// Mitsubishi GX Works2 project: 11国轩烘烤线体修改1028   PLC: Q06UDEH

TYPE ConveyorIO : STRUCT
  xUnloadCCW : BOOL;  (* 下料为反转 *)
  xUnloadAlarm : BOOL;  (* 下料报警 *)
  xUnload : BOOL;  (* 下料请求 *)
  xPutInto : BOOL;  (* 线体直接投入物料 *)
  xNotArriveAlarm : BOOL;  (* 未到达报警 *)
  xNextRun : BOOL;  (* 下段线体运行 *)
  xMotorCW : BOOL;  (* 电机正转 *)
  xMotorCCW : BOOL;  (* 电机反转 *)
  xManual : BOOL;  (* 手动 *)
  xloadCCW : BOOL;  (* 上料为反转 *)
  xLimitAlarrm : BOOL;  (* 限位报警 *)
  xLoad : BOOL;  (* 上料请求 *)
  xForward : BOOL;  (* 正转手动 *)
  xEmpty : BOOL;  (* 线体状态为空 *)
  xCWPresent : BOOL;  (* 正转检测有无传感器 *)
  xCCWPresent : BOOL;  (* 反转检测有无传感器 *)
  xBusy : BOOL;  (* 工作中 *)
  xBackward : BOOL;  (* 反转手动 *)
  xAuto : BOOL;  (* 自动 *)
  xPosLimit : BOOL;  (* 正限位 *)
  xNegLimit : BOOL;  (* 负限位 *)
  xOverWidthAlarm : BOOL;  (* 超宽报警 *)
  xError : BOOL;  (* 报警 *)
  iProductCategoryIn : INT;  (* 产品类型输入 *)
  iProductCategory : INT;  (* 产品类型记录 *)
  iProductCategoryOut : INT;  (* 产品类型输出 *)
  diDeviceID : DINT;  (* 设备编号 *)
  tUnloadAlarmDelay : TIME;  (* 下料报警时间设置 *)
  tLoadDelay : TIME;  (* 上料延时设置 *)
  xSizeDeficientDetect : BOOL;  (* 尺寸缺陷检测 *)
  xZoneClear : BOOL;  (* 初始化线体清除 *)
  tZoneClearTime : TIME;  (* 初始化线体清除时间 *)
  iTaskIDIn : INT;  (* 产品类型输入 *)
  iTaskID : INT;  (* 产品类型记录 *)
  iTaskIDOut : INT;  (* 产品类型输出 *)
  diDesConveyorIn : DINT;  (* 产品类型输入 *)
  diDesConveyor : DINT;  (* 产品类型记录 *)
  diDesConveyorOut : DINT;  (* 产品类型输出 *)
END_STRUCT END_TYPE

TYPE ShuttleCarIO : STRUCT
  xReady : BOOL;  (* 准备就绪 *)
  xForward : BOOL;  (* 正转 *)
  xBackward : BOOL;  (* 反转 *)
  iCurrentPos : INT;  (* 当前位置 *)
  iDestinationPos : INT;  (* 目标位置 *)
  xCW : BOOL;  (* 正转输出 *)
  xCCW : BOOL;  (* 反转输出 *)
  xBrake : BOOL;  (* 刹车 *)
  xHomeSwitch : BOOL;  (* 零位接近开关 *)
  xPosLimit : BOOL;  (* 正限位 *)
  xNegLimit : BOOL;  (* 负限位 *)
  xMDIExe : BOOL;  (* MDI开始 *)
  xMDIDone : BOOL;  (* MDI 完成 *)
  xPassLimit : BOOL;  (* 限位屏蔽 *)
  xPosLimitCatch : BOOL;  (* 正限位捕捉 *)
  xNegLimitCatch : BOOL;  (* 负限位捕捉 *)
  xHomeExe : BOOL;  (* 开始寻零 *)
  xHomeDone : BOOL;  (* 寻零完成 *)
  xHomeBusy : BOOL;  (* 寻零中 *)
  xHomeFailed : BOOL;  (* 寻零失败 *)
  xBusy : BOOL;  (* 工作中 *)
  tArriveDelay : TIME;  (* 到位延时 *)
  xCylinder : BOOL;  (* 气缸控制 *)
  tBrakeDelay : TIME;  (* 抱闸延时 *)
  xPauseRamp : BOOL;  (* 暂停减速斜坡标志位 *)
  xPresentDetect1 : BOOL;  (* 物料有无检测1 *)
  xPresentDetect2 : BOOL;  (* 物料有无检测2 *)
  xOvertimeAlarm : BOOL;  (* 超时报警 *)
  tSetOverTime : TIME;  (* 设置超时时间 *)
  xLooseDetect : BOOL;  (* 松绳检测 *)
  xLooseAlarm : BOOL;  (* 松绳报警 *)
  xArrive : BOOL;  (* 到位信号 *)
  diDeviceID : DINT;  (* 设备编号 *)
  xMoveStep : BOOL;  (* 寸动 *)
  xAdrSwitch : ARRAY [1..8] OF BOOL;  (* 位置开关 *)
END_STRUCT END_TYPE

TYPE SwitchIO : STRUCT
  xLiftCylinderRetractDetect : BOOL;
  xLiftCylinderExtendDetect : BOOL;
  xLiftCylinderRetract : BOOL;
  xLiftCylinderExtend : BOOL;
  xEntryBarCylinderRetract : BOOL;
  xLiftCylinderExtendInit : BOOL;
  xEntryEnable : BOOL;
  xExitEnable : BOOL;
  xExitBarCylinderRetract : BOOL;
  xSwithEnable : BOOL;
  xLiftCylinderRetractButton : BOOL;
  xLiftCylinderExtendButton : BOOL;
  xEntryBarCylinderRetractButton : BOOL;
  xExitBarCylinderRetractButton : BOOL;
  xPutInto : BOOL;  (* 单体复位 *)
  tSetOvertime : TIME;  (* 设定超时报警时间 *)
  xOvertimeAlarm : BOOL;  (* 超时报警 *)
END_STRUCT END_TYPE

TYPE QueueElement : STRUCT
  xCondition : BOOL;
  iPriority : INT;
END_STRUCT END_TYPE

TYPE UConveyorIO : STRUCT
  xLiftCylinderRetractDetect1 : BOOL;  (* 左臂顶升移栽收回检测 *)
  xLiftCylinderRetractDetect2 : BOOL;  (* 右臂顶升移栽收回检测 *)
  xLiftCylinderExtendDetect1 : BOOL;  (* 左臂顶升移栽顶起检测 *)
  xLiftCylinderExtendDetect2 : BOOL;  (* 右臂顶升移栽顶起检测 *)
  xLiftCylinderRetract1 : BOOL;  (* 左臂顶升移栽收回输出1 *)
  xLiftCylinderRetract2 : BOOL;  (* 右臂顶升移栽收回输出2 *)
  xLiftCylinderExtend1 : BOOL;  (* 左臂顶升移栽顶起输出1 *)
  xLiftCylinderExtend2 : BOOL;  (* 右臂顶升移栽顶起输出2 *)
  xExitBarCylinderRetract1 : BOOL;  (* 左臂阻挡收回输出1 *)
  xExitBarCylinderRetract2 : BOOL;  (* 右臂阻挡收回输出2 *)
  xLiftCylinderExtendInit1 : BOOL;  (* 左臂顶升移栽初始状态 *)
  xLiftCylinderExtendInit2 : BOOL;  (* 右臂顶升移栽初始状态 *)
  xEntryEnable1 : BOOL;  (* U型1线体入使能 *)
  xEntryEnable2 : BOOL;  (* U型2线体入使能 *)
  xEntryEnable3 : BOOL;  (* U型3线体入使能 *)
  xExitEnable1 : BOOL;  (* U型1线体出使能 *)
  xExitEnable2 : BOOL;  (* U型2线体出使能 *)
  xExitEnable3 : BOOL;  (* U型3线体出使能 *)
  xPassEnable : BOOL;  (* 直接放行去下段 *)
  xLiftCylinderRetractButton1 : BOOL;  (* 顶升移栽收回按钮1 *)
  xLiftCylinderRetractButton2 : BOOL;  (* 顶升移栽收回按钮2 *)
  xLiftCylinderExtendButton1 : BOOL;  (* 顶升移栽顶起按钮1 *)
  xLiftCylinderExtendButton2 : BOOL;  (* 顶升移栽顶起按钮2 *)
  xExitBarCylinderRetractButton1 : BOOL;  (* 阻挡气缸1 *)
  xExitBarCylinderRetractButton2 : BOOL;  (* 阻挡气缸2 *)
  xPutInto : BOOL;  (* 单体复位 *)
  tSetOvertime : TIME;  (* 设定超时报警时间 *)
  xOvertimeAlarm : BOOL;  (* 超时报警 *)
  iTask : INT;  (* 3个任务执行步骤 *)
  xBatteryDetect1 : BOOL;  (* 电池检测1 *)
  xBatteryDetect2 : BOOL;  (* 电池检测2 *)
  xBatteryError : BOOL;  (* 空框检测到电池报警 *)
END_STRUCT END_TYPE

TYPE CommunicationIO : STRUCT
  i_iResponsPCPLC : INT;  (* 上位机写入-请求确认 *)
  i_iReadWriteFlagPCPLC : INT;  (* 上位机写入-读写标志位 *)
  i_iTaskProcessFlagPCPLC : INT;  (* 上位机写入-任务出料标志位 *)
  i_iCommandPCPLC : INT;  (* 上位机写入-命令字 *)
  i_iTaskIDPCPLC : INT;  (* 上位机写入-任务号 *)
  i_diDestinationDevicePCPLC : DINT;  (* 上位机写入-目标设备号 *)
  i_iProductIDPCPLC : INT;  (* 上位机写入-框码后4位 *)
  o_iRequestPLCPC : INT;  (* 上位机读取-请求状态 *)
  o_iReadWriteFlagPLCPC : INT;  (* 上位机读取-读写标志位 *)
  o_iDeviceStatusPLCPC : INT;  (* 上位机读取-设备状态 *)
  o_iTaskIDPLCPC : INT;  (* 上位机读取-任务号 *)
  o_iProductIDPLCPC : INT;  (* 上位机读取-框码后4位 *)
END_STRUCT END_TYPE

// global labels: Global
VAR_GLOBAL
  g_xTcpFailed : BOOL;
  g_xPickOver : ARRAY [1..4] OF BOOL;  (* 注液机给我们的信号，待定 *)
  g_xPickStart : ARRAY [1..4] OF BOOL;  (* 我们给注液机信号，开始挑选 *)
  m_lky1 AT M25 : BOOL;
  m_xLoadPermit1 AT M52 : BOOL;  (* 允许生成上料任务(可触摸屏，也可自动) *)
  m_xLoadPermit3 AT M54 : BOOL;  (* 允许生成上料任务(可触摸屏，也可自动) *)
  m_xLoadPermit2 AT M53 : BOOL;  (* 允许生成上料任务(可触摸屏，也可自动) *)
  m_xLoadPermit4 AT M55 : BOOL;  (* 允许生成上料任务(可触摸屏，也可自动) *)
  m_xLoadPermit5 AT M56 : BOOL;  (* 允许生成上料任务(可触摸屏，也可自动) *)
  g_xAuto AT M11 : BOOL;
  g_xAutoSwitch AT X1 : BOOL;
  g_xManual : BOOL;
  g_xEStop AT X0 : BOOL;
  g_xReset AT X4 : BOOL;
  g_xResetSingle AT M4 : BOOL;  (* 单线体复位 *)
  g_xInsertTask AT M5 : BOOL;  (* 插入任务 *)
  g_iInsertTaskID AT D2 : INT;  (* 插入任务号 *)
  g_iInsertCategory AT D6 : INT;
  g_diInsertDesConveyor AT D8 : DINT;
  g_iConveyorStatus AT D4 : INT;
  g_xAlarm : BOOL;
  g_xMute AT M15 : BOOL;
  g_xStackLampRed AT Y200 : BOOL;
  g_xStackLampAmber AT Y201 : BOOL;
  g_xStackLampGreen AT Y202 : BOOL;
  g_xBuzzer AT Y203 : BOOL;
  g_xStop AT X3 : BOOL;
  g_xPause AT M3 : BOOL;  (* 暂停 *)
  g_xAutoStart AT X2 : BOOL;
  g_xAutoLamp AT Y204 : BOOL;
  g_xRemoteAutoStart AT M0 : BOOL;
  g_xRemoteAuto AT M10 : BOOL;
  g_iState AT D40 : INT;
  g_iLocalAutoStep : BOOL;
  g_diDeviceIDSelect AT D0 : DINT;
END_VAR

// task Task_01 (event TRUE, interval 0, priority 31): POU, TCP, start

PROGRAM POU
VAR
  Conveyor11102 : Conveyor;
  Conveyor11104 : Conveyor;
  Conveyor11105 : Conveyor;
  Conveyor11106 : Conveyor;
  Conveyor11103 : Conveyor;
  Conveyor11107 : Conveyor;
  Conveyor11108 : Conveyor;
  Conveyor11101 : Conveyor;
  Conveyor11109 : Conveyor;
  Conveyor11110 : Conveyor;
  Conveyor11111 : Conveyor;
  Conveyor11112 : Conveyor;
  Conveyor11113 : Conveyor;
  Conveyor11114 : Conveyor;
  Conveyor11115 : Conveyor;
  Conveyor11116 : Conveyor;
  Conveyor11117 : Conveyor;
  Conveyor11118 : Conveyor;
  Conveyor111181 : Conveyor;
  Conveyor11119 : Conveyor;
  Conveyor11120 : Conveyor;
  Conveyor111201 : Conveyor;
  Conveyor11121 : Conveyor;
  Conveyor111211 : Conveyor;
  Conveyor11122 : Conveyor;
  Conveyor11123 : Conveyor;
  Conveyor111231 : Conveyor;
  Conveyor11124 : Conveyor;
  Conveyor111241 : Conveyor;
  Conveyor11125 : Conveyor;
  Conveyor11126 : Conveyor;
  Conveyor111261 : Conveyor;
  Conveyor11127 : Conveyor;
  Conveyor111271 : Conveyor;
  Conveyor11128 : Conveyor;
  Conveyor11129 : Conveyor;
  Conveyor111291 : Conveyor;
  Conveyor11130 : Conveyor;
  Conveyor11131 : Conveyor;
  Conveyor11132 : Conveyor;
  Conveyor11133 : Conveyor;
  Conveyor11134 : Conveyor;
  Conveyor11135 : Conveyor;
  Conveyor11136 : Conveyor;
  Conveyor11137 : Conveyor;
  Conveyor11138 : Conveyor;
  Conveyor11139 : Conveyor;
  Conveyor11140 : Conveyor;
  Conveyor11141 : Conveyor;
  Conveyor11142 : Conveyor;
  Conveyor11143 : Conveyor;
  Conveyor11144 : Conveyor;
  ConveyorIO11101 : ConveyorIO;
  ConveyorIO11102 : ConveyorIO;
  ConveyorIO11103 : ConveyorIO;
  ConveyorIO11104 : ConveyorIO;
  ConveyorIO11105 : ConveyorIO;
  ConveyorIO11106 : ConveyorIO;
  ConveyorIO11107 : ConveyorIO;
  ConveyorIO11108 : ConveyorIO;
  ConveyorIO11109 : ConveyorIO;
  ConveyorIO11110 : ConveyorIO;
  ConveyorIO11111 : ConveyorIO;
  ConveyorIO11112 : ConveyorIO;
  ConveyorIO11113 : ConveyorIO;
  ConveyorIO11114 : ConveyorIO;
  ConveyorIO11115 : ConveyorIO;
  ConveyorIO11116 : ConveyorIO;
  ConveyorIO11117 : ConveyorIO;
  ConveyorIO11118 : ConveyorIO;
  ConveyorIO111181 : ConveyorIO;
  ConveyorIO11119 : ConveyorIO;
  ConveyorIO11120 : ConveyorIO;
  ConveyorIO111201 : ConveyorIO;
  ConveyorIO11121 : ConveyorIO;
  ConveyorIO111211 : ConveyorIO;
  ConveyorIO11122 : ConveyorIO;
  ConveyorIO11123 : ConveyorIO;
  ConveyorIO111231 : ConveyorIO;
  ConveyorIO11124 : ConveyorIO;
  ConveyorIO111241 : ConveyorIO;
  ConveyorIO11125 : ConveyorIO;
  ConveyorIO11126 : ConveyorIO;
  ConveyorIO111261 : ConveyorIO;
  ConveyorIO11127 : ConveyorIO;
  ConveyorIO111271 : ConveyorIO;
  ConveyorIO11128 : ConveyorIO;
  ConveyorIO11129 : ConveyorIO;
  ConveyorIO111291 : ConveyorIO;
  ConveyorIO11130 : ConveyorIO;
  ConveyorIO11131 : ConveyorIO;
  ConveyorIO11132 : ConveyorIO;
  ConveyorIO11133 : ConveyorIO;
  ConveyorIO11134 : ConveyorIO;
  ConveyorIO11135 : ConveyorIO;
  ConveyorIO11136 : ConveyorIO;
  ConveyorIO11137 : ConveyorIO;
  ConveyorIO11138 : ConveyorIO;
  ConveyorIO11139 : ConveyorIO;
  ConveyorIO11140 : ConveyorIO;
  ConveyorIO11141 : ConveyorIO;
  ConveyorIO11142 : ConveyorIO;
  ConveyorIO11143 : ConveyorIO;
  ConveyorIO11144 : ConveyorIO;
  Lifter11202 : ShuttleCar;  (* 烘烤去注液口升降机 *)
  Lifter11203 : ShuttleCar;  (* 注液回流升降机 *)
  LifterIO11202 : ShuttleCarIO;  (* 烘烤去注液口升降机 *)
  LifterIO11203 : ShuttleCarIO;  (* 注液回流升降机 *)
  Switch11301 : Switch;  (* 上层交叉点 *)
  Switch11302 : Switch;  (* 烘烤入库 *)
  UConveyor11303 : UConveyor;  (* 注液1 *)
  UConveyor11306 : UConveyor;  (* 注液2 *)
  UConveyor11309 : UConveyor;  (* 注液3 *)
  UConveyor11312 : UConveyor;  (* 注液4 *)
  UConveyorIO11303 : UConveyorIO;  (* 注液1 *)
  UConveyorIO11306 : UConveyorIO;  (* 注液2 *)
  UConveyorIO11309 : UConveyorIO;  (* 注液3 *)
  UConveyorIO11312 : UConveyorIO;  (* 注液4 *)
  Switch11301Task : PreemptivePriority;  (* 上层交叉点抢栈任务 *)
  Switch11301Condition : ARRAY [1..13] OF BOOL;  (* 上层交叉点抢栈任务 *)
  m_i11301Task : INT;  (* 上层交叉点抢栈任务 *)
  Switch11316Task : PriorityQueue;  (* 下层出库排队任务 *)
  Switch11316Condition : ARRAY [1..13] OF QueueElement;  (* 下层出库排队任务 *)
  m_i11316Task : INT;  (* 下层出库排队任务 *)
  Switch11315Task : PreemptivePriority;  (* 下层交叉点抢栈任务 *)
  Switch11315Condition : ARRAY [1..13] OF BOOL;  (* 下层交叉点抢栈任务 *)
  Conveyor11139Task : PriorityQueue;  (* 注液入排队任务 *)
  Conveyor11139Condition : ARRAY [1..13] OF QueueElement;  (* 注液入排队任务 *)
  m_i11139Task : INT;  (* 注液入排队任务 *)
  m_xPickDone : ARRAY [1..4] OF BOOL;  (* 他给信号，我们自己置位一个信号 *)
  Uconveyor11303Task : PreemptivePriority;  (* 注液1任务 *)
  Uconveyor11303Condition : ARRAY [1..13] OF BOOL;  (* 注液1条件 *)
  Uconveyor11306Task : PreemptivePriority;  (* 注液2任务 *)
  Uconveyor11306Condition : ARRAY [1..13] OF BOOL;  (* 注液2条件 *)
  Uconveyor11309Task : PreemptivePriority;  (* 注液3任务 *)
  Uconveyor11309Condition : ARRAY [1..13] OF BOOL;  (* 注液3条件 *)
  Uconveyor11312Task : PreemptivePriority;  (* 注液4任务 *)
  Uconveyor11312Condition : ARRAY [1..13] OF BOOL;  (* 注液4条件 *)
  Cylinder11304 : ShuttleCar;  (* 注液处顶升1 *)
  Cylinder11307 : ShuttleCar;  (* 注液处顶升2 *)
  Cylinder11310 : ShuttleCar;  (* 注液处顶升3 *)
  Cylinder11313 : ShuttleCar;  (* 注液处顶升4 *)
  Cylinder112011 : ShuttleCar;  (* 上层门升降1 *)
  Cylinder112012 : ShuttleCar;  (* 上层门升降2 *)
  Cylinder112041 : ShuttleCar;  (* 下层门升降1 *)
  Cylinder112042 : ShuttleCar;  (* 下层门升降2 *)
  CylinderIO11304 : ShuttleCarIO;  (* 注液处顶升1 *)
  CylinderIO11307 : ShuttleCarIO;  (* 注液处顶升2 *)
  CylinderIO11310 : ShuttleCarIO;  (* 注液处顶升3 *)
  CylinderIO11313 : ShuttleCarIO;  (* 注液处顶升4 *)
  CylinderIO112011 : ShuttleCarIO;  (* 上层门升降1 *)
  CylinderIO112012 : ShuttleCarIO;  (* 上层门升降2 *)
  CylinderIO112041 : ShuttleCarIO;  (* 下层门升降1 *)
  CylinderIO112042 : ShuttleCarIO;  (* 下层门升降2 *)
  m_xLoadPermit : ARRAY [1..4] OF BOOL;  (* 允许生成上料任务(可触摸屏，也可自动) *)
  ComConveyor11104 : ConveyorCommunication;  (* 烘烤入库扫码 *)
  ComConveyor11108 : ConveyorCommunication;  (* 烘烤1入库有料 *)
  ComConveyor11107 : ConveyorCommunication;  (* 烘烤2入库有料 *)
  ComConveyor11142 : ConveyorCommunication;  (* 烘烤1出库完成 *)
  ComConveyor11141 : ConveyorCommunication;  (* 烘烤2出库完成 *)
  ComConveyor11110 : ConveyorCommunication;  (* 品检区 *)
  ComConveyor11111 : ConveyorCommunication;  (* 注液前扫码 *)
  ComConveyor11143 : ConveyorCommunication;  (* 烘烤后入组装 *)
  ComConveyorIO11104 : CommunicationIO;  (* 烘烤入库扫码 *)
  ComConveyorIO11108 : CommunicationIO;  (* 烘烤1入库有料 *)
  ComConveyorIO11107 : CommunicationIO;  (* 烘烤2入库有料 *)
  ComConveyorIO11142 : CommunicationIO;  (* 烘烤1出库完成 *)
  ComConveyorIO11141 : CommunicationIO;  (* 烘烤2出库完成 *)
  ComConveyorIO11110 : CommunicationIO;  (* 品检区 *)
  ComConveyorIO11111 : CommunicationIO;  (* 注液前扫码 *)
  ComConveyorIO11143 : CommunicationIO;  (* 烘烤后入组装 *)
  m_i11315Task : INT;  (* 下层交叉点抢栈任务 *)
  Switch11315 : Switch;  (* 烘烤出库 *)
  Switch11316 : Switch;  (* 下层交叉点 *)
  SwitchIO11301 : SwitchIO;  (* 上层交叉点 *)
  SwitchIO11302 : SwitchIO;  (* 烘烤入库 *)
  SwitchIO11315 : SwitchIO;  (* 烘烤出库 *)
  SwitchIO11316 : SwitchIO;  (* 下层交叉点 *)
  Conveyor11145 : Conveyor;
  Conveyor11146 : Conveyor;
  Conveyor11147 : Conveyor;
  ConveyorIO11145 : ConveyorIO;
  ConveyorIO11146 : ConveyorIO;
  ConveyorIO11147 : ConveyorIO;
  m_Ton315 : TON;
  m_x315 : BOOL;  (* 315顶升移栽检测延时 *)
  m_t315 : TIME;
  Conveyor111381 : Conveyor;
  ConveyorIO111381 : ConveyorIO;
  ConveyorIO111382 : ConveyorIO;
  Conveyor111382 : Conveyor;
  ConveyorIO111041 : ConveyorIO;
  Conveyor111041 : Conveyor;
  Conveyor111042 : Conveyor;
  ConveyorIO111042 : ConveyorIO;
  m_TPU1TaskComplete : TP;  (* U1完成延时 *)
  m_tU1TaskComplete : TIME;  (* U1完成延时 *)
  m_xU1TaskComplete : BOOL;  (* U1完成延时 *)
  m_TPU2TaskComplete : TP;  (* U2完成延时 *)
  m_tU2TaskComplete : TIME;  (* U2完成延时 *)
  m_xU2TaskComplete : BOOL;  (* U2完成延时 *)
  m_TPU3TaskComplete : TP;  (* U3完成延时 *)
  m_tU3TaskComplete : TIME;  (* U3完成延时 *)
  m_xU3TaskComplete : BOOL;  (* U3完成延时 *)
  m_TPU4TaskComplete : TP;  (* U4完成延时 *)
  m_tU4TaskComplete : TIME;  (* U4完成延时 *)
  m_xU4TaskComplete : BOOL;  (* U4完成延时 *)
  m_TonU1TaskStart : TON;  (* U1任务开始延时 *)
  m_tU1TaskStart : TIME;  (* U1任务开始延时 *)
  m_xU1TaskStart : BOOL;  (* U1任务开始延时 *)
  m_TonU2TaskStart : TON;  (* U2任务开始延时 *)
  m_tU2TaskStart : TIME;  (* U2任务开始延时 *)
  m_xU2TaskStart : BOOL;  (* U2任务开始延时 *)
  m_TonU3TaskStart : TON;  (* U3任务开始延时 *)
  m_tU3TaskStart : TIME;  (* U3任务开始延时 *)
  m_xU3TaskStart : BOOL;  (* U3任务开始延时 *)
  m_TonU4TaskStart : TON;  (* U4任务开始延时 *)
  m_tU4TaskStart : TIME;  (* U4任务开始延时 *)
  m_xU4TaskStart : BOOL;  (* U4任务开始延时 *)
  m_Ton11119 : TON;  (* 11119有料延时刷新111201定时器 *)
  m_t111201 : TIME;  (* 111201延时计时 *)
  m_x111201 : BOOL;  (* 111201延时刷新 *)
  ConveyorIO111315Entry : ConveyorIO;
  ConveyorIO111315Exit : ConveyorIO;
  Conveyor111315Entry : Conveyor;
  Conveyor111315Exit : Conveyor;
  m_Ton11122 : TON;  (* 11122有料延时刷新111211定时器 *)
  m_t111211 : TIME;  (* 111211延时计时 *)
  m_x111211 : BOOL;  (* 111211延时刷新 *)
  m_Ton11125 : TON;  (* 11125有料延时刷新111261定时器 *)
  m_t111261 : TIME;  (* 111261延时计时 *)
  m_x111261 : BOOL;  (* 111261延时刷新 *)
  Lifter11204 : ShuttleCar;  (* 烘烤出库1顶升气缸 *)
  Lifter11205 : ShuttleCar;  (* 烘烤出库2顶升气缸 *)
  LifterIO11204 : ShuttleCarIO;  (* 烘烤出库1顶升气缸 *)
  LifterIO11205 : ShuttleCarIO;  (* 烘烤出库2顶升气缸 *)
  m_11119communication : BOOL;  (* 与机械手对接信号标志位1 *)
  m_11122communication : BOOL;  (* 与机械手对接信号标志位2 *)
  m_11125communication : BOOL;  (* 与机械手对接信号标志位3 *)
  m_11128communication : BOOL;  (* 与机械手对接信号标志位4 *)
  m_Ton11128 : TON;  (* 11128有料延时刷新111271定时器 *)
  m_t111271 : TIME;  (* 111271延时计时 *)
  m_x111271 : BOOL;  (* 111271延时刷新 *)
  m_Ton11141 : TON;  (* 11141有料延时刷新定时器 *)
  m_t11141 : TIME;  (* 11141延时计时 *)
  m_x11141 : BOOL;  (* 11141延时刷新 *)
END_VAR
 
Conveyor11101(ConveyorMotor:=	ConveyorIO11101);
ConveyorIO11101.xCWPresent:=X08;
Y208:=ConveyorIO11101.xMotorCW;
ConveyorIO11101.xForward:=M500;
M301:=NOT ConveyorIO11101.xEmpty;
F401:=ConveyorIO11101.xUnloadAlarm;
ConveyorIO11101.diDeviceID:=11101;
ConveyorIO11101.tLoadDelay:=T#1S;

Conveyor11102(ConveyorMotor:=	ConveyorIO11102);
ConveyorIO11102.xCWPresent:=X9;
Y209:=ConveyorIO11102.xMotorCW;
ConveyorIO11102.xForward:=M501;
M302:=NOT ConveyorIO11102.xEmpty;
F402:=ConveyorIO11102.xUnloadAlarm;
ConveyorIO11102.diDeviceID:=11102;


Conveyor11103(ConveyorMotor:=	ConveyorIO11103);
ConveyorIO11103.xCWPresent:=XA;
M303:=NOT ConveyorIO11103.xEmpty;
F403:=ConveyorIO11103.xUnloadAlarm;
Y20A:=ConveyorIO11103.xMotorCW;
ConveyorIO11103.xForward:=M502;
ConveyorIO11103.diDeviceID:=11103;
ConveyorIO11103.tLoadDelay:=T#4S;

Conveyor11104(ConveyorMotor:=	ConveyorIO11104);
ConveyorIO11104.xCWPresent:=XB;
Y20B:=ConveyorIO11104.xMotorCW OR ConveyorIO111041.xMotorCW;
ConveyorIO11104.xForward:=M503;
M304:=NOT ConveyorIO11104.xEmpty;
F404:=ConveyorIO11104.xUnloadAlarm;
ConveyorIO11104.diDeviceID:=11104;

Conveyor111041(ConveyorMotor:=	ConveyorIO111041);
ConveyorIO111041.xCWPresent:=XA;
ConveyorIO111041.diDeviceID:=111041;
ConveyorIO111041.tLoadDelay:=T#5S;


Conveyor111042(ConveyorMotor:=	ConveyorIO111042);
ConveyorIO111042.xCWPresent:=XC;
ConveyorIO111042.diDeviceID:=111042;
ConveyorIO111042.tLoadDelay:=T#8S;

Conveyor11105(ConveyorMotor:=	ConveyorIO11105);
ConveyorIO11105.xCWPresent:=X16;
Y238:=ConveyorIO11105.xMotorCW;
ConveyorIO11105.xForward:=M504;
M305:=NOT ConveyorIO11105.xEmpty;
F405:=ConveyorIO11105.xUnloadAlarm;
ConveyorIO11105.diDeviceID:=11105;

Conveyor11106(ConveyorMotor:=	ConveyorIO11106);
ConveyorIO11106.xCWPresent:=XC;
Y20D:=ConveyorIO11106.xMotorCW;
ConveyorIO11106.xForward:=M505;
Y20E:=ConveyorIO11106.xMotorCCW;					
ConveyorIO11106.xBackward:=M506;					
M306:=NOT ConveyorIO11106.xEmpty;
F406:=ConveyorIO11106.xUnloadAlarm;
ConveyorIO11106.diDeviceID:=11106;

Conveyor11107(ConveyorMotor:=	ConveyorIO11107);
ConveyorIO11107.xCWPresent:=XE;
Y20F:=ConveyorIO11107.xMotorCW;
ConveyorIO11107.xForward:=M507;
M307:=NOT ConveyorIO11107.xEmpty;
F407:=ConveyorIO11107.xUnloadAlarm;
ConveyorIO11107.diDeviceID:=11107;
ConveyorIO11107.tLoadDelay:=T#3s;
ConveyorIO11107.xPutInto:=SM412;

Conveyor11108(ConveyorMotor:=	ConveyorIO11108);
ConveyorIO11108.xCWPresent:=XF;
Y210:=ConveyorIO11108.xMotorCW;
ConveyorIO11108.xForward:=M508;
M308:=NOT ConveyorIO11108.xEmpty;
F408:=ConveyorIO11108.xUnloadAlarm;
ConveyorIO11108.diDeviceID:=11108;
ConveyorIO11108.tLoadDelay:=T#3S;

Conveyor11109(ConveyorMotor:=	ConveyorIO11109);
ConveyorIO11109.xCWPresent:=X10;	(*需根据正转方向修改*)
ConveyorIO11109.xCCWPresent:=X11;	
ConveyorIO11109.xNegLimit:=NOT X12;				
Y211:=ConveyorIO11109.xMotorCW;	
Y212:=ConveyorIO11109.xMotorCCW;					
ConveyorIO11109.xForward:=M509;	
ConveyorIO11109.xBackward:=M510;					
M309:=NOT ConveyorIO11109.xEmpty;
F409:=ConveyorIO11109.xUnloadAlarm;
ConveyorIO11109.diDeviceID:=11109;

Conveyor11110(ConveyorMotor:=	ConveyorIO11110);
ConveyorIO11110.xCWPresent:=X14;(*需修改*)
ConveyorIO11110.xNegLimit:=X15;		
Y213:=ConveyorIO11110.xMotorCW;
ConveyorIO11110.xForward:=M511;			
M310:=NOT ConveyorIO11110.xEmpty;
F410:=ConveyorIO11110.xUnloadAlarm;
ConveyorIO11110.diDeviceID:=11110;

Conveyor11111(ConveyorMotor:=	ConveyorIO11111);
ConveyorIO11111.xCWPresent:=X58;
Y214:=ConveyorIO11111.xMotorCW;
ConveyorIO11111.xForward:=M512;	
M311:=NOT ConveyorIO11111.xEmpty;
F411:=ConveyorIO11111.xUnloadAlarm;
ConveyorIO11111.diDeviceID:=11111;


Conveyor11112(ConveyorMotor:=	ConveyorIO11112);
ConveyorIO11112.xCWPresent:=X59;
Y215:=ConveyorIO11112.xMotorCW;
ConveyorIO11112.xForward:=M513;
M313:=NOT ConveyorIO11112.xEmpty;
F413:=ConveyorIO11112.xUnloadAlarm;
ConveyorIO11112.diDeviceID:=11112;

Conveyor11113(ConveyorMotor:=	ConveyorIO11113);
Y216:=ConveyorIO11113.xMotorCW;
ConveyorIO11113.xForward:=M514;
M314:=NOT ConveyorIO11113.xEmpty;
F414:=ConveyorIO11113.xUnloadAlarm;
ConveyorIO11113.diDeviceID:=11113;
ConveyorIO11113.tLoadDelay:=T#2S;

Conveyor11114(ConveyorMotor:=	ConveyorIO11114);
Y217:=ConveyorIO11114.xMotorCW;
ConveyorIO11114.xForward:=M515;
M315:=NOT ConveyorIO11114.xEmpty;
F415:=ConveyorIO11114.xUnloadAlarm;
ConveyorIO11114.diDeviceID:=11114;
ConveyorIO11114.tLoadDelay:=T#2S;

Conveyor11115(ConveyorMotor:=	ConveyorIO11115);
Y218:=ConveyorIO11115.xMotorCW;
ConveyorIO11115.xForward:=M516;
M316:=NOT ConveyorIO11115.xEmpty;
F416:=ConveyorIO11115.xUnloadAlarm;
ConveyorIO11115.diDeviceID:=11115;
ConveyorIO11115.tLoadDelay:=T#2S;

Conveyor11116(ConveyorMotor:=	ConveyorIO11116);
ConveyorIO11116.xPosLimit:=NOT X28;
Y219:=ConveyorIO11116.xMotorCW;
ConveyorIO11116.xForward:=M517;
M317:=NOT ConveyorIO11116.xEmpty;
F417:=ConveyorIO11116.xUnloadAlarm;
ConveyorIO11116.diDeviceID:=11116;
ConveyorIO11116.tLoadDelay:=T#2S;

Conveyor11117(ConveyorMotor:=	ConveyorIO11117);
ConveyorIO11117.xCWPresent:=X2A;(*根据正转方向更改*)
ConveyorIO11117.xNegLimit:=NOT X29;
Y21A:=ConveyorIO11117.xMotorCW;
ConveyorIO11117.xForward:=M518;					
Y21B:=ConveyorIO11117.xMotorCCW;					
ConveyorIO11117.xBackward:=M519;					
M318:=NOT ConveyorIO11117.xEmpty;
F418:=ConveyorIO11117.xUnloadAlarm;
ConveyorIO11117.diDeviceID:=11117;

Conveyor11118(ConveyorMotor:=	ConveyorIO11118);
ConveyorIO11118.xCCWPresent:=X1B;
Y21C:=ConveyorIO11118.xMotorCW;
ConveyorIO11118.xForward:=M520;
M319:=NOT ConveyorIO111181.xEmpty;
F419:=ConveyorIO11118.xUnloadAlarm;
ConveyorIO11118.diDeviceID:=11118;
ConveyorIO11118.tLoadDelay:=T#5S;

Conveyor111181(ConveyorMotor:=	ConveyorIO111181);
ConveyorIO111181.xCWPresent:=X2C;
ConveyorIO111181.diDeviceID:=111181;
ConveyorIO111181.tLoadDelay:=T#11S;

Conveyor11119(ConveyorMotor:=	ConveyorIO11119);
ConveyorIO11119.xCWPresent:=X2D;
Y21D:=ConveyorIO11119.xMotorCW;
ConveyorIO11119.xForward:=M521;
M321:=NOT ConveyorIO11119.xEmpty;
F421:=ConveyorIO11119.xUnloadAlarm;
ConveyorIO11119.diDeviceID:=11119;
ConveyorIO11119.tLoadDelay:=T#3S;

Conveyor11120(ConveyorMotor:=	ConveyorIO11120);
ConveyorIO11120.xCWPresent:=X19;
Y21E:=ConveyorIO11120.xMotorCCW;
ConveyorIO11120.xBackward:=M522;
M322:=NOT ConveyorIO111201.xEmpty;
F422:=ConveyorIO111201.xUnloadAlarm;
ConveyorIO11120.diDeviceID:=11120;
ConveyorIO11120.tLoadDelay:=T#8S;

Conveyor111201(ConveyorMotor:=	ConveyorIO111201);
ConveyorIO111201.xCWPresent:=X2D;
ConveyorIO111201.diDeviceID:=1111201;

Conveyor11121(ConveyorMotor:=	ConveyorIO11121);
ConveyorIO11121.xCCWPresent:=X1C;
Y21F:=ConveyorIO11121.xMotorCCW;
ConveyorIO11121.xloadCCW:=1;
ConveyorIO11121.xBackward:=M523;
M324:=NOT ConveyorIO111211.xEmpty;
F424:=ConveyorIO11121.xUnloadAlarm;
ConveyorIO11121.diDeviceID:=11121;
ConveyorIO11121.tLoadDelay:=T#3S;

Conveyor111211(ConveyorMotor:=	ConveyorIO111211);
ConveyorIO111211.xCWPresent:=X30;
ConveyorIO111211.diDeviceID:=1111211;

Conveyor11122(ConveyorMotor:=	ConveyorIO11122);
ConveyorIO11122.xCWPresent:=X30;
Y23D:=ConveyorIO11122.xMotorCW;
ConveyorIO11122.xForward:=M524;
M326:=NOT ConveyorIO11122.xEmpty;
F426:=ConveyorIO11122.xUnloadAlarm;
ConveyorIO11122.diDeviceID:=11122;
ConveyorIO11122.tLoadDelay:=T#2S;

Conveyor11123(ConveyorMotor:=	ConveyorIO11123);
ConveyorIO11123.xCcWPresent:=X1D;
Y221:=ConveyorIO11123.xMotorCW;
ConveyorIO11123.xForward:=M525;
M327:=NOT ConveyorIO111231.xEmpty;
F427:=ConveyorIO111231.xUnloadAlarm;
ConveyorIO11123.diDeviceID:=11123;

Conveyor111231(ConveyorMotor:=	ConveyorIO111231);
ConveyorIO111231.xCWPresent:=X31;
ConveyorIO111231.diDeviceID:=111231;
ConveyorIO111231.tLoadDelay:=T#11S;

Conveyor11124(ConveyorMotor:=	ConveyorIO11124);
ConveyorIO11124.xCCWPresent:=X20;
M329:=NOT ConveyorIO111241.xEmpty;
F429:=ConveyorIO11124.xUnloadAlarm;
ConveyorIO11124.diDeviceID:=11124;

Conveyor111241(ConveyorMotor:=	ConveyorIO111241);
ConveyorIO111241.xCWPresent:=X32;
Y222:=ConveyorIO111241.xMotorCW;
ConveyorIO111241.xForward:=M526;
ConveyorIO111241.diDeviceID:=111241;
ConveyorIO111241.tLoadDelay:=T#5S;

Conveyor11125(ConveyorMotor:=	ConveyorIO11125);
ConveyorIO11125.xCWPresent:=X33;
Y223:=ConveyorIO11125.xMotorCW;
ConveyorIO11125.xForward:=M527;
ConveyorIO11125.diDeviceID:=11125;
ConveyorIO11125.tLoadDelay:=T#2S;

Conveyor11126(ConveyorMotor:=	ConveyorIO11126);
ConveyorIO11126.xCCWPresent:=X21;
Y224:=ConveyorIO11126.xMotorCCW;
ConveyorIO11126.xBackward:=M528;
M332:=NOT ConveyorIO111261.xEmpty;
F432:=ConveyorIO111261.xUnloadAlarm;
ConveyorIO11126.diDeviceID:=11126;
ConveyorIO11126.tLoadDelay:=T#3S;

Conveyor111261(ConveyorMotor:=	ConveyorIO111261);
ConveyorIO111261.xCWPresent:=X33;
ConveyorIO111261.diDeviceID:=1111261;

Conveyor11127(ConveyorMotor:=	ConveyorIO11127);
ConveyorIO11127.xCCWPresent:=X24;
Y225:=ConveyorIO11127.xMotorCCW;
ConveyorIO11127.xBackward:=M529;
M334:=NOT ConveyorIO111271.xEmpty;
F434:=ConveyorIO11127.xUnloadAlarm;
ConveyorIO11127.diDeviceID:=11127;
ConveyorIO11127.tLoadDelay:=T#3S;

Conveyor111271(ConveyorMotor:=	ConveyorIO111271);
ConveyorIO111271.xCWPresent:=X36;
ConveyorIO111271.diDeviceID:=1111271;

Conveyor11128(ConveyorMotor:=	ConveyorIO11128);
ConveyorIO11128.xCWPresent:=X36;
Y226:=ConveyorIO11128.xMotorCW;
ConveyorIO11128.xForward:=M530;
M336:=NOT ConveyorIO11128.xEmpty;
F436:=ConveyorIO11128.xUnloadAlarm;
ConveyorIO11128.diDeviceID:=11128;
ConveyorIO11128.tLoadDelay:=T#2S;


Conveyor11129(ConveyorMotor:=	ConveyorIO11129);
ConveyorIO11129.xCCWPresent:=X25;
Y227:=ConveyorIO11129.xMotorCW;
ConveyorIO11129.xForward:=M531;
M337:=NOT ConveyorIO111291.xEmpty;
F437:=ConveyorIO111291.xUnloadAlarm;
ConveyorIO11129.diDeviceID:=11129;

Conveyor111291(ConveyorMotor:=	ConveyorIO111291);
ConveyorIO111291.xCWPresent:=X37;
ConveyorIO111291.diDeviceID:=111291;
ConveyorIO111291.tLoadDelay:=T#5S;

Conveyor11130(ConveyorMotor:=	ConveyorIO11130);
ConveyorIO11130.xCWPresent:=X38;
Y228:=ConveyorIO11130.xMotorCW;
ConveyorIO11130.xForward:=M532;
M339:=NOT ConveyorIO11130.xEmpty;
F439:=ConveyorIO11130.xUnloadAlarm;
ConveyorIO11130.diDeviceID:=11130;

Conveyor11131(ConveyorMotor:=	ConveyorIO11131);
ConveyorIO11131.xCWPresent:=X39;
Y229:=ConveyorIO11131.xMotorCW;
ConveyorIO11131.xForward:=M533;
M340:=NOT ConveyorIO11131.xEmpty;
F440:=ConveyorIO11131.xUnloadAlarm;
ConveyorIO11131.diDeviceID:=11131;

Conveyor11132(ConveyorMotor:=	ConveyorIO11132);
ConveyorIO11132.xCWPresent:=X3A;
Y22A:=ConveyorIO11132.xMotorCW;
ConveyorIO11132.xForward:=M534;
M341:=NOT ConveyorIO11132.xEmpty;
F441:=ConveyorIO11132.xUnloadAlarm;
ConveyorIO11132.diDeviceID:=11132;

Conveyor11133(ConveyorMotor:=	ConveyorIO11133);
ConveyorIO11133.xCWPresent:=X3B;
Y22B:=ConveyorIO11133.xMotorCW;
ConveyorIO11133.xForward:=M535;
M342:=NOT ConveyorIO11133.xEmpty;
F442:=ConveyorIO11133.xUnloadAlarm;
ConveyorIO11133.diDeviceID:=11133;

Conveyor11134(ConveyorMotor:=	ConveyorIO11134);
ConveyorIO11134.xCWPresent:=X3C;
Y22C:=ConveyorIO11134.xMotorCW;
ConveyorIO11134.xForward:=M536;
M343:=NOT ConveyorIO11134.xEmpty;
F443:=ConveyorIO11134.xUnloadAlarm;
ConveyorIO11134.diDeviceID:=11134;

Conveyor11135(ConveyorMotor:=	ConveyorIO11135);
ConveyorIO11135.xCWPresent:=X3D;
Y22D:=ConveyorIO11135.xMotorCW;
ConveyorIO11135.xForward:=M537;
M344:=NOT ConveyorIO11135.xEmpty;
F444:=ConveyorIO11135.xUnloadAlarm;
ConveyorIO11135.diDeviceID:=11135;

Conveyor11136(ConveyorMotor:=	ConveyorIO11136);
ConveyorIO11136.xCWPresent:=X3E;
Y22E:=ConveyorIO11136.xMotorCW;
ConveyorIO11136.xForward:=M538;
M345:=NOT ConveyorIO11136.xEmpty;
F445:=ConveyorIO11136.xUnloadAlarm;
ConveyorIO11136.diDeviceID:=11136;

Conveyor11137(ConveyorMotor:=	ConveyorIO11137);
ConveyorIO11137.xCWPresent:=X41;
Y22F:=ConveyorIO11137.xMotorCW;
ConveyorIO11137.xForward:=M539;
M346:=NOT ConveyorIO11137.xEmpty;
F446:=ConveyorIO11137.xUnloadAlarm;
ConveyorIO11137.diDeviceID:=11137;
ConveyorIO11137.tLoadDelay:=T#4S;

Conveyor11138(ConveyorMotor:=	ConveyorIO11138);
ConveyorIO11138.xCWPresent:=X43;
Y230:=ConveyorIO11138.xMotorCW OR ConveyorIO111381.xMotorCW OR ConveyorIO111382.xMotorCW;
ConveyorIO11138.xForward:=M540;
M347:=NOT ConveyorIO11138.xEmpty;
F447:=ConveyorIO11138.xUnloadAlarm;
ConveyorIO11138.diDeviceID:=11138;

Conveyor111381(ConveyorMotor:=	ConveyorIO111381);
ConveyorIO111381.xCWPresent:=X41;
ConveyorIO11138.diDeviceID:=11138;
ConveyorIO111381.tLoadDelay:=T#5S;

Conveyor111382(ConveyorMotor:=	ConveyorIO111382);
ConveyorIO111382.xCWPresent:=X44;
ConveyorIO111382.diDeviceID:=11138;
ConveyorIO111382.tLoadDelay:=T#5S;

Conveyor11139(ConveyorMotor:=	ConveyorIO11139);
ConveyorIO11139.xCWPresent:=X17;
Y239:=ConveyorIO11139.xMotorCW;
ConveyorIO11139.xForward:=M541;
M348:=NOT ConveyorIO11139.xEmpty;
F448:=ConveyorIO11139.xUnloadAlarm;
ConveyorIO11139.diDeviceID:=11139;

Conveyor11140(ConveyorMotor:=	ConveyorIO11140);
ConveyorIO11140.xCWPresent:=X44;
Y232:=ConveyorIO11140.xMotorCW;
Y233:=ConveyorIO11140.xMotorCCW;
ConveyorIO11140.xForward:=M542;
ConveyorIO11140.xBackward:=M543;
M349:=NOT ConveyorIO11140.xEmpty;
F449:=ConveyorIO11140.xUnloadAlarm;
ConveyorIO11140.diDeviceID:=11140;
ConveyorIO11140.tLoadDelay:=T#5S;

Conveyor11141(ConveyorMotor:=	ConveyorIO11141);
ConveyorIO11141.xCWPresent:=X46;
Y234:=ConveyorIO11141.xMotorCW;
ConveyorIO11141.xForward:=M544;
M350:=NOT ConveyorIO11141.xEmpty;
F450:=ConveyorIO11141.xUnloadAlarm;
ConveyorIO11141.diDeviceID:=11141;
m_Ton11141(IN:=X46,
					PT:=T#30s,
					Q:= m_x11141,
					ET:=m_t11141);
ConveyorIO11141.xPutInto:=m_x11141;


Conveyor11142(ConveyorMotor:=	ConveyorIO11142);
ConveyorIO11142.xCWPresent:=X47;
Y235:=ConveyorIO11142.xMotorCW;
ConveyorIO11142.xForward:=M545;
M351:=NOT ConveyorIO11142.xEmpty;
F451:=ConveyorIO11142.xUnloadAlarm;
ConveyorIO11142.diDeviceID:=11142;

Conveyor11143(ConveyorMotor:=	ConveyorIO11143);
ConveyorIO11143.xCWPresent:=X49;
ConveyorIO11143.xCCWPresent:=X49;
Y236:=ConveyorIO11143.xMotorCW;
ConveyorIO11143.xForward:=M546;
M352:=NOT ConveyorIO11143.xEmpty;
F452:=ConveyorIO11143.xUnloadAlarm;
ConveyorIO11143.diDeviceID:=11143;

Conveyor11144(ConveyorMotor:=	ConveyorIO11144);
ConveyorIO11144.xCWPresent:=X48;
Y237:=ConveyorIO11144.xMotorCW;
ConveyorIO11144.xForward:=M547;
M353:=NOT ConveyorIO11144.xEmpty;
F453:=ConveyorIO11144.xUnloadAlarm;
ConveyorIO11144.diDeviceID:=11144;
ConveyorIO11144.tLoadDelay:=T#1S;

(*新增上层3段线体*)
Conveyor11145(ConveyorMotor:=	ConveyorIO11145);
ConveyorIO11145.xCWPresent:=X5A(*根据现场接线修改*);
Y23A:=ConveyorIO11145.xMotorCW;
ConveyorIO11145.xForward:=M588(*根据现场接线修改*);
M354:=NOT ConveyorIO11145.xEmpty;
F454:=ConveyorIO11145.xUnloadAlarm;
ConveyorIO11145.diDeviceID:=11145;

Conveyor11146(ConveyorMotor:=	ConveyorIO11146);
ConveyorIO11146.xCWPresent:=X5B;
Y23B:=ConveyorIO11146.xMotorCW;
ConveyorIO11146.xForward:=M589(*根据现场接线修改*);
M355:=NOT ConveyorIO11146.xEmpty;
F455:=ConveyorIO11146.xUnloadAlarm;
ConveyorIO11146.diDeviceID:=11146;


Conveyor11147(ConveyorMotor:=	ConveyorIO11147);
ConveyorIO11147.xCWPresent:=X5C;
Y23C:=ConveyorIO11147.xMotorCW;
ConveyorIO11147.xForward:=M590(*根据现场接线修改*);
M356:=NOT ConveyorIO11147.xEmpty;
F456:=ConveyorIO11147.xUnloadAlarm;
ConveyorIO11147.diDeviceID:=11147;



(*————————————————————————————————————————————————*)

Lifter11202(ShuttleCarInOut:=LifterIO11202);(*入口侧升降台*)
LifterIO11202.xCylinder:=1;
Y244:=LifterIO11202.xCW;(*修改*)	
Y245:=LifterIO11202.xCCW;(*修改*)	
LifterIO11202.xForward:=M548;
LifterIO11202.xBackward:=M549;
ShuttleCarCurrentPosition(X4F OR X4E,X4E,X4F,FALSE,LifterIO11202.iCurrentPos);
F454:=LifterIO11202.xOvertimeAlarm ;
LifterIO11202.diDeviceID:=11202;

lifter11203(ShuttleCarInOut:=LifterIO11203);(*出口升降台*)
LifterIO11203.xCylinder:=1;
Y246:=LifterIO11203.xCW;
Y247:=LifterIO11203.xCCW;
LifterIO11203.xForward:=M550;
LifterIO11203.xBackward:=M551;
ShuttleCarCurrentPosition(X51 OR X50,X50,X51,FALSE,LifterIO11203.iCurrentPos);
F455:=LifterIO11203.xOvertimeAlarm ;
LifterIO11203.diDeviceID:=11203;
(*烘烤出库下层线体新增2个顶升气缸*)
lifter11204(ShuttleCarInOut:=LifterIO11204);(*烘烤1出口升降台*)
LifterIO11204.xCylinder:=1;
Y26A:=LifterIO11204.xCW;
Y26B:=LifterIO11204.xCCW;
LifterIO11204.xForward:=M725;(*需修改*)
LifterIO11204.xBackward:=M724;(*需修改*)
ShuttleCarCurrentPosition(X81 OR X80,X81,X80,FALSE,LifterIO11204.iCurrentPos);
F455:=LifterIO11204.xOvertimeAlarm ;(*需修改*)
LifterIO11204.diDeviceID:=11204;(*需修改*)

lifter11205(ShuttleCarInOut:=LifterIO11205);(*烘烤2出口升降台*)
LifterIO11205.xCylinder:=1;
Y26C:=LifterIO11205.xCW;
Y26D:=LifterIO11205.xCCW;
LifterIO11205.xForward:=M726;(*需修改*)
LifterIO11205.xBackward:=M727;(*需修改*)
ShuttleCarCurrentPosition(X82 OR X83,X82,X83,FALSE,LifterIO11205.iCurrentPos);
F455:=LifterIO11205.xOvertimeAlarm ;(*需修改*)
LifterIO11205.diDeviceID:=11205;(*需修改*)